(* CODESYS project Revisora(2)_V3_0_2k.project
   Company: Schneider Electric
   Title: Revisora
   Author: Frank Willian
   Version: 2.0.0.0

Project tree, tasks and I/O mapping:
  MyController : TM241CE40T/U, Schneider Electric, order no. TM241CE40T/U, version 4.0.6.18
    application Application
      libraries: SysTime, 3.4.1.20 (System)
      task MAST (cyclic, interval 10 ms, priority 15, watchdog 100 ms x 1) calls R00_main
      task Task1ms (cyclic, interval 1 ms, priority 1) calls RB01_enableReb
      global variables GVL
      01_Maquina/
        program R06_principal [LD]
        program R01_firstScan [LD]
        program R05_comando [LD]
        program R20_acessorios [LD]
        program R99_calcTempos [ST]
        program R00_main [LD]
        program R30_receita [ST]
        program R19_cilindros [LD]
        program R18_alinhador [LD]
        program R50_reset [ST]
      Structs/
        data type _exec_bits
        data type _eixo_drive
        data type _eixo_home
        data type _eixo_auto
        data type _receita
        data type _eixo
      05_IHM/
        program I02_alarmes [ST]
        program I06_textoConfirma [LD]
        program I01_geral [LD]
        program I03_mensagens [ST]
      03_Nip/
        program NP03_auto [LD]
        program NP01_geral [LD]
        program NP06_jog [LD]
        program NP09_sentido [ST]
        program NP04_parada [LD]
        program NP02_enableNip [LD]
        program NP07_veloc [ST]
        program NP20_JogTest [ST]
      global variables PersistentVars
      global variables IHM
      Symbol configuration
      Visu/
      10_Relogio/
        function block GetDateAndTime [CFC]
        function block SetDateAndTime [CFC]
        program AjustaDataHora [LD]
      image pool Imagens
      11_FB/
        function block RTO [ST]
      02_Rebobinadores/
        program RB01_enableReb [LD]
        program RB05_sentido [ST]
        program RB03_analog [LD]
        program RB04_saidas [LD]
      19_Ultra/
        program U10_auto [LD]
    Cartridge_1 : Cartridge, Schneider Electric, version 4.0.6.18
    Cartridge_2 : Cartridge, Schneider Electric, version 4.0.6.18
    IO_Bus : IO bus - TM3, Schneider Electric, version 4.0.6.18
      Saidas_Analog : TM3AQ2/G, Schneider Electric, order no. TM3AQ2/G, version 1.0.0.12
          settings: KPI Configuration.KPI Configuration[0] = 17; KPI Configuration.KPI Configuration[1] = 17; KPI Configuration.KPI Configuration[2] = 240; KPI Configuration.KPI Configuration[3] = 216; KPI Configuration.KPI Configuration[4] = 240; KPI Configuration.KPI Configuration[5] = 216; KPI Configuration.KPI Configuration[6] = 16; KPI Configuration.KPI Configuration[7] = 39; KPI Configuration.KPI Configuration[8] = 16; KPI Configuration.KPI Configuration[9] = 39
          output analoReb01 : INT  // QW0
          output analoReb02 : INT  // QW1
          input  ibAnalog_IBStatusQW0 : BYTE  // IBStatusQW0
          input  ibAnalog_IBStatusQW1 : BYTE  // IBStatusQW1
      Entradas_Analog : TM3AI4/G, Schneider Electric, order no. TM3AI4/G, version 1.0.0.15
          settings: KPI Configuration.KPI Configuration[0] = 34; KPI Configuration.KPI Configuration[1] = 34; KPI Configuration.KPI Configuration[5] = 0; KPI Configuration.KPI Configuration[7] = 0; KPI Configuration.KPI Configuration[12] = 32; KPI Configuration.KPI Configuration[13] = 78; KPI Configuration.KPI Configuration[14] = 32; KPI Configuration.KPI Configuration[15] = 78
          input  ia_sensorUltraSom_1 : INT  // IW0
          input  ia_sensorUltraSom_2 : INT  // IW1
          input  iiModule_1_IW2 : INT  // IW2
          input  iiModule_1_IW3 : INT  // IW3
          input  ibModule_1_IBStatusIW0 : BYTE  // IBStatusIW0
          input  ibModule_1_IBStatusIW1 : BYTE  // IBStatusIW1
          input  ibModule_1_IBStatusIW2 : BYTE  // IBStatusIW2
          input  ibModule_1_IBStatusIW3 : BYTE  // IBStatusIW3
    COM_Bus : COM bus, Schneider Electric, version 4.0.6.18
    Ethernet_1 : Ethernet Network, Schneider Electric, version 4.0.6.18
        settings: IPAddress = [192, 168, 1, 10]; SubnetMask = [255, 255, 255, 0]; WebServer = TRUE; FTP Server = TRUE; SoMachine Protocol = TRUE; Modbus Server = TRUE; NetManage Protocol = TRUE; SNMP protocol = TRUE; WebVisu protocol = TRUE
    Serial_Line_1 : Serial line, Schneider Electric, version 4.0.6.18
      SoMachine_Network_Manager : SoMachine-Network Manager, Schneider Electric, version 4.0.0.2
    Serial_Line_2 : Serial line, Schneider Electric, version 4.0.6.18
      Modbus_Manager : Modbus Manager, Schneider Electric, version 4.0.0.2
    DI : Digital Inputs, Schneider Electric, version 4.0.6.18
        input  i_releEmergencia : BOOL  // IDW0.I0
        input  i_btReset : BOOL  // IDW0.I1
        input  i_ligaRevisora : BOOL  // IDW0.I2
        input  i_sentido : BOOL  // IDW0.I4
        input  i_cortina : BOOL  // IDW0.I6
        input  i_finalDeContagem : BOOL  // IDW0.I9
        unmapped channels: IDW0, IB1
    DQ : Digital Outputs, Schneider Electric, version 4.0.6.18
        settings: Outputs Usage = 15
        output o_enableReb01 : BOOL  // QW0.Q4
        output o_enableNip : BOOL  // QW0.Q5
        output o_enableReb02 : BOOL  // QW0.Q6
        output o_alinhador : BOOL  // QW0.Q7
        output o_mesaCentro : BOOL  // QW0.Q8
        output o_cilindroNip : BOOL  // QW0.Q9
        output o_mesaAuto : BOOL  // QW0.Q10
        output o_abilitaPulsoNip : BOOL  // QW0.Q11
        output qbDQ_QB1 : BYTE  // QB1
        unmapped channels: QW0
    Counters : Counters, Schneider Electric, version 4.0.6.18
    Pulse_Generators : Pulse Generators, Schneider Electric, version 4.0.6.18
        settings: Instance name = 'nip_PTO'; B output History = 'old=-1 new=1'; A output History = 'old=-1 new=0'; Temporary Instance name = 'nip_PTO'; Instance name = 'selag_PTO'; B output History = 'old=-1 new=3'; A output History = 'old=-1 new=2'; Temporary Instance name = 'selag_PTO'
  HMISTU855 : HMIS5T, Schneider Electric, order no. HMIS5T, version 3.5.3.54
    HMI Application
    Ethernet
      SoMachine_Network_Manager2 : SoMachine-Network Manager, Schneider Electric, version 4.0.0.2
    USB
      SoMachine_Network_Manager3 : SoMachine-Network Manager, Schneider Electric, version 4.0.0.2
    COM1
      SoMachine_Network_Manager1 : SoMachine-Network Manager, Schneider Electric, version 4.0.0.2
  6c0f7fb6-600b-4c93-9262-20cdc603757e
  text list GlobalTextList
  5ce3da45-db07-42e7-a21c-a00fff4ed8f6|C:\_Clientes\Opuspac\Doc\Figuras\Botao.png
  5ce3da45-db07-42e7-a21c-a00fff4ed8f6|C:\_Clientes\Opuspac\Doc\Figuras\Botao_ps.png
  5ce3da45-db07-42e7-a21c-a00fff4ed8f6|C:\_Clientes\Opuspac\Doc\Figuras\LogoOpus.jpg
  Vijeo Designer Project Container
*)

// MyController/Application/Structs/_exec_bits
TYPE _exec_bits :
STRUCT
	RQ					: BOOL;
	IP					: BOOL;
	DN					: BOOL;
	Fase				: DINT;
	Mask				: DINT;
END_STRUCT
END_TYPE

// MyController/Application/Structs/_eixo_drive
TYPE _eixo_drive :
STRUCT
	falha			: MC_ReadAxisError_PTO;
	posicao			: MC_ReadActualPosition_PTO;
	power			: MC_Power_PTO;
	reset			: MC_Reset_PTO;
	state			: MC_ReadMotionState_PTO;
	status			: MC_ReadStatus_PTO;
	stop			: MC_Stop_PTO;
END_STRUCT
END_TYPE

// MyController/Application/Structs/_eixo_home
TYPE _eixo_home :
STRUCT
	RQ					: BOOL;
	IP					: BOOL;
	DN					: BOOL;
	Fase				: DINT;
	Mask				: DINT;
	movVeloc			: MC_MoveVelocity_PTO;
	movRelat			: MC_MoveRelative_PTO;
	movStop				: ARRAY[1..2] OF MC_Stop_PTO;
	setPos				: MC_SetPosition_PTO;
END_STRUCT
END_TYPE

// MyController/Application/Structs/_eixo_auto
TYPE _eixo_auto :
STRUCT
	movVeloc					: ARRAY [1..3] OF MC_MoveVelocity_PTO;
	movAbs						: MC_MoveAbsolute_PTO;
	movRelat					: ARRAY [0..3] OF MC_MoveRelative_PTO;
	movStop						: MC_Stop_PTO;
	setPos						: MC_SetPosition_PTO;
END_STRUCT
END_TYPE

// MyController/Application/Structs/_receita
TYPE _receita :
STRUCT
	
	velocDesb		: DINT;
	velocReb		: DINT;
	freioDesb		: INT;
	freioReb		: INT;
	torqueDesb		: INT;
	torqueReb		: INT;

END_STRUCT
END_TYPE

// MyController/Application/Structs/_eixo
TYPE _eixo :
STRUCT
	auto				: _eixo_auto;
	home				: _eixo_home;
	drive				: _eixo_drive;
	falha				: BOOL;
	posicaoAtual		: DINT;
	calcula				: BOOL;
	parando				: BOOL;
	pausa				: BOOL;
	constMove			: BOOL;
	errorStop			: BOOL;
END_STRUCT
END_TYPE

// MyController/Application/GVL
VAR_GLOBAL
	
	jogNip						: BOOL;
	jogRebEsq					: BOOL;
	jogRebDir					: BOOL;
	jogDirecao					: BOOL;
	jogAbilita					: BOOL;
	jogEnebleGeral				: BOOL;
	jogCilindroNip				: BOOL;
	valorPorcRebobinador		: ARRAY [1..2] OF REAL;
	tempoAtrasoAposDesligar		: BOOL;
	troggerTest					: BOOL;
	cortinaOk					: BOOL;
	mudaVeloc					: BOOL;
	auxAnaloReb01				: INT;
	auxAnaloReb02				: INT;
	abilitaTrocaVeloc			: BOOL;
	abilitaPulsoNip				: _exec_bits;
	T_desabilitaPulsoNip		: TON;
	tpoDesabilitaPulsoNip		: BOOL;
	
	
	// transições
	psBtCiclo					: BOOL;

	// Variaveis gerais
	alarmeReset					: BOOL;
	alarmeResetInd				: BOOL;
	alwaysOff					: BOOL;
	alwaysOn					: BOOL;
	calcGeral					: BOOL;
	calcTempos					: BOOL;
	comandoOff					: BOOL;
	emergOk						: BOOL;
	existeAlarme				: BOOL;
	firstScan					: BOOL;
	injecaoTpoOff				: BOOL;
	ladoDir						: BOOL;
	ladoEsq						: BOOL;
	liberaCiclo					: BOOL;
	ligaAlinhador				: BOOL;
	livreComando				: BOOL;
	livreStart					: BOOL;
	ligaMaq						: BOOL;
	manual						: BOOL;
	mesaCentro					: BOOL;
	modoAutomatico				: BOOL;
	nipEmMove					: BOOL;
	nipPausado					: BOOL;
	partidaOK					: BOOL;
	partidaLenta				: BOOL;
	velocPartida				: BOOL;		
	pisca						: BOOL;
	piscaRapido					: BOOL;
	primeiroCiclo				: BOOL;
	start						: BOOL;
	sentidoDesbobinar			: BOOL;
	sentidoRebobinar			: BOOL;
	torqueParada				: BOOL;
	triggerBobina				: BOOL;
	triggerValorDesbReb			: BOOL;
	
	tpoInicio					: TIME;
	
	revisora					: _eixo;
	nip							: _eixo;

	TL_inicializa				: TON;
	T_nipLiga					: TON;
	
	alinhador					: _exec_bits;
	ciclo						: _exec_bits;
	contagem					: _exec_bits;
	cilNip						: _exec_bits;
	comando						: _exec_bits;
	enbReb						: _exec_bits;
	enbNip						: _exec_bits;
	liga						: _exec_bits;
	desliga						: _exec_bits;
	jogNeg						: _exec_bits;
	jogPos						: _exec_bits;
	nipMove						: _exec_bits;
	nipParada					: _exec_bits;
	nipStop						: _exec_bits;
	principal					: _exec_bits;	


	porcRebobinador				: ARRAY [1..2] OF REAL;
	rebobiPorc 					: ARRAY [1..2] OF LIN_TRAFO;
	
    //Sincroniza e ajusta o relógio da IHM
	AnoSet						: UINT;
	ClkScan						: BOOL;
	AjustaHora					: BOOL;
	MesSet						: UINT;
	DiaSet						: UINT;
	HoraSet						: UINT;
	MinutoSet					: UINT;
	SegundoSet					: UINT;
	AnoAtual					: UINT;
	MesAtual					: UINT;
	DiaAtual					: UINT;
	HoraAtual					: UINT;
	MinutoAtual					: UINT;
	SegundoAtual				: UINT;	
	sink						: BOOL;

(*	=================== ALARMES ===================
	Obs: alarme[0]- Não utilizado
*)
	alarme						: ARRAY[0..50] OF BOOL;
	alarmes						: _exec_bits;
	mensagem					: ARRAY[0..50] OF BOOL;
	numAlarme					: SINT;
		
(*	=================== Alterações ===================  *)
	ativoManual					: BOOL;
	tpoArAtivo					: TIME;

(*	=================== Ultrassonico ===================  *)	
	rebobTorqueOper				: ARRAY[0..2] OF REAL;
	desbobTorqueOper			: ARRAY[0..2] OF REAL;
	analogTorqueDrive			: ARRAY[0..2] OF INT;


END_VAR

// MyController/Application/PersistentVars
VAR_GLOBAL PERSISTENT RETAIN
	versaoSoftware				: REAL:= 1.00;
	pi							: REAL:= 3.1415926;
	paramFab					: BOOL:= TRUE;
	numRec						: SINT;
	displayState				: INT;
	jogVelocNip					: DINT;
	revisoraVelocNip			: DINT;
	valorJogRebob01				: INT;
	valorJogRebob02				: INT;
		
	// NIP
	auxVeloc					: ARRAY[0..4] OF BOOL;
	saidaReb					: ARRAY[0..1] OF BOOL;
	M_diamRolo					: DINT:= 34;
	M_revisoraVeloc				: DINT;
	M_revisoraAcel				: DINT:= 800;
	M_revisoraDecel				: DINT:= 200;
	M_pulsosParar				: DINT;
	parseAnalog					: ARRAY[0..1] OF INT;
	ihm_velocidade				: DINT:= 10;
	ihm_tempoInicio				: DINT:= 10;
	visLadoDir					: BOOL;
	visLadoEsq					: BOOL;
	
	veloc						: ARRAY[0..4] OF DINT;
	delayTorq					: ARRAY[0..1] OF TIME;
	sentido						: INT;
	
	bobina			 			: ARRAY[0..5] OF _receita;	
	bobinaAtual					: _receita;
	
	//	========= ultrassonico ===========	
	ihm_btUltraSomHab			: BOOL;
	
	//	========= desbobinador ===========	
	M_desbobTorqueMin				: ARRAY[0..2] OF REAL;
	M_desbobTorqueMax				: ARRAY[0..2] OF REAL;
	M_desbobTorqueOper				: ARRAY[0..2] OF REAL;
	valorDesbobTorqueMin			: REAL;
	valorDesbobTorqueMax			: REAL;
	
	//  ========== Rebobinador ===========
	M_rebobTorqueMin				: ARRAY[0..2] OF REAL;
	M_rebobTorqueMax				: ARRAY[0..2] OF REAL;
	M_rebobTorqueOper				: ARRAY[0..2] OF REAL;
	valorRebobTorqueMin				: REAL;
	valorRebobTorqueMax				: REAL;

END_VAR

// MyController/Application/IHM
VAR_GLOBAL
	ihm_alarme					: ARRAY[0..50] OF BOOL;
	ihm_alarmeReset				: BOOL;
	ihm_alarmeResetInd			: BOOL;
	ihm_bannerConfirma			: BOOL;
	ihm_bannerMensagem			: BOOL;
	ihm_confirmaV				: BOOL;
	ihm_confirmaX				: BOOL;
	ihm_mensagem				: DINT;
	ihm_numReceita				: SINT;
	ihm_telaHome				: BOOL;
	ihm_telaAtual				: INT;
	ihm_textoConfirma			: DINT;
	ihm_textoProced				: DINT;
	ihm_velocMedida				: DINT;
	ihm_inverte					: BOOL;
	ihm_cilindroNip				: BOOL;
	ihm_alinhador				: BOOL;
	nome						: WSTRING;
	
	ihm_valorDesb				: ARRAY[0..2] OF REAL;
	ihm_valorReb				: ARRAY[0..2] OF REAL;
	
	ihm_desbobInc				: BOOL;
	ihm_desbobDec				: BOOL;
	
	ihm_rebobInc				: BOOL;
	ihm_rebobDec				: BOOL;

END_VAR

// MyController/Application/01_Maquina/R00_main
PROGRAM R00_main
VAR
END_VAR

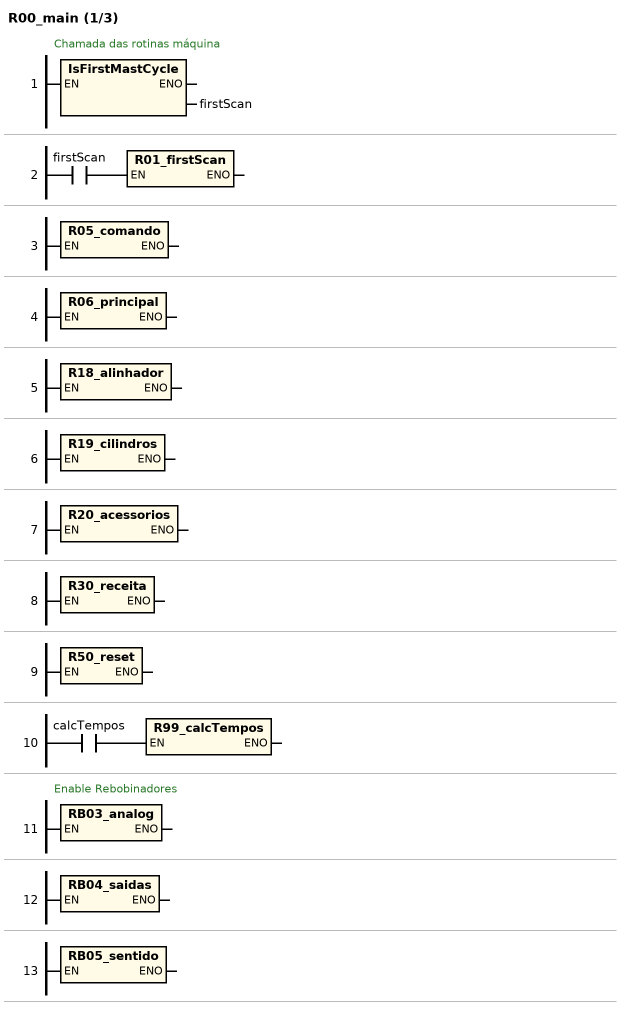
// NETWORK 1
// Chamada das rotinas máquina
firstScan := IsFirstMastCycle();

// NETWORK 2
IF firstScan THEN R01_firstScan(); END_IF

// NETWORK 3
R05_comando();

// NETWORK 4
R06_principal();

// NETWORK 5
R18_alinhador();

// NETWORK 6
R19_cilindros();

// NETWORK 7
R20_acessorios();

// NETWORK 8
R30_receita();

// NETWORK 9
R50_reset();

// NETWORK 10
IF calcTempos THEN R99_calcTempos(); END_IF

// NETWORK 11
// Enable Rebobinadores
RB03_analog();

// NETWORK 12
RB04_saidas();

// NETWORK 13
RB05_sentido();

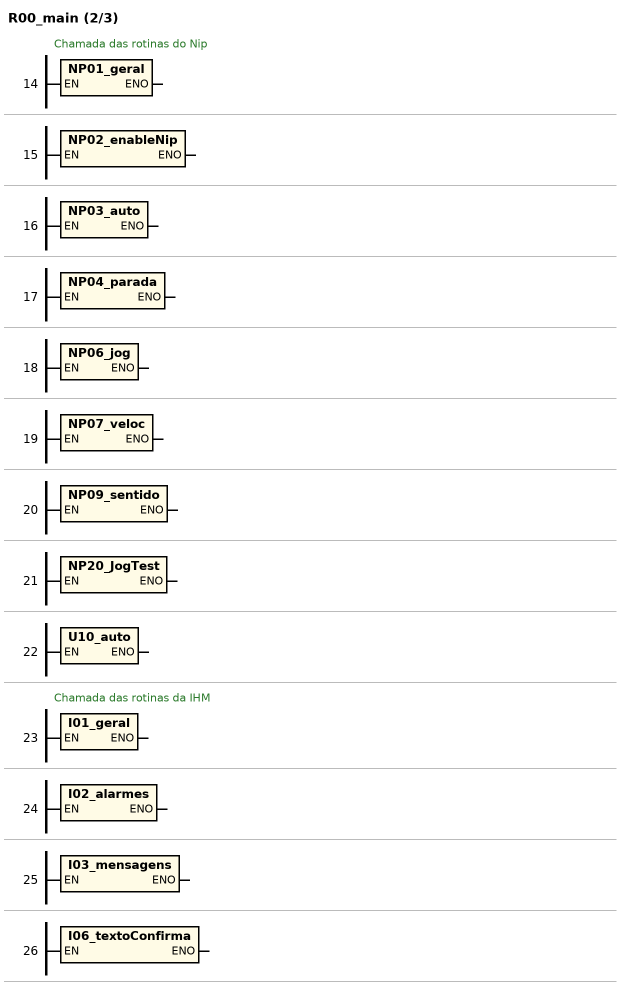
// NETWORK 14
// Chamada das rotinas do Nip
NP01_geral();

// NETWORK 15
NP02_enableNip();

// NETWORK 16
NP03_auto();

// NETWORK 17
NP04_parada();

// NETWORK 18
NP06_jog();

// NETWORK 19
NP07_veloc();

// NETWORK 20
NP09_sentido();

// NETWORK 21
NP20_JogTest();

// NETWORK 22
U10_auto();

// NETWORK 23
// Chamada das rotinas da IHM
I01_geral();

// NETWORK 24
I02_alarmes();

// NETWORK 25
I03_mensagens();

// NETWORK 26
I06_textoConfirma();

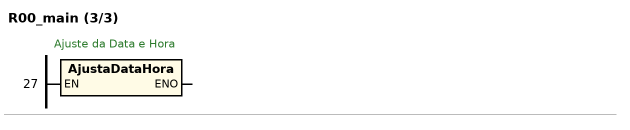
// NETWORK 27
// Ajuste da Data e Hora
AjustaDataHora();

END_PROGRAM

// MyController/Application/01_Maquina/R01_firstScan
PROGRAM R01_firstScan
VAR
END_VAR

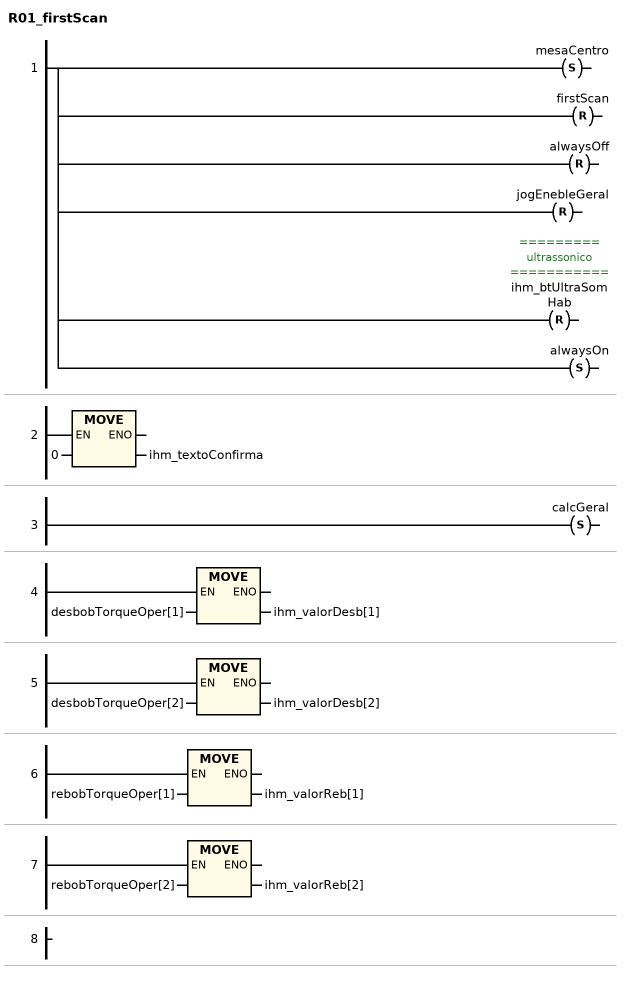
// NETWORK 1
//   ihm_btUltraSomHab: ========= ultrassonico ===========
mesaCentro S= TRUE;
firstScan R= TRUE;
alwaysOff R= TRUE;
jogEnebleGeral R= TRUE;
ihm_btUltraSomHab R= TRUE;
alwaysOn S= TRUE;

// NETWORK 2
ihm_textoConfirma := 0;

// NETWORK 3
calcGeral S= TRUE;

// NETWORK 4
ihm_valorDesb[1] := desbobTorqueOper[1];

// NETWORK 5
ihm_valorDesb[2] := desbobTorqueOper[2];

// NETWORK 6
//   rebobTorqueOper[1]: =================== Ultrassonico ===================
ihm_valorReb[1] := rebobTorqueOper[1];

// NETWORK 7
//   rebobTorqueOper[2]: =================== Ultrassonico ===================
ihm_valorReb[2] := rebobTorqueOper[2];

// NETWORK 8

END_PROGRAM

// MyController/Application/01_Maquina/R05_comando
PROGRAM R05_comando
VAR
	TL_comando				: TON;
END_VAR
VAR // added by the converter: edge detectors and wires of the graphical bodies
    _rt1 : R_TRIG;
    _ft1, _ft2 : F_TRIG;
    _w1 : BOOL;
END_VAR

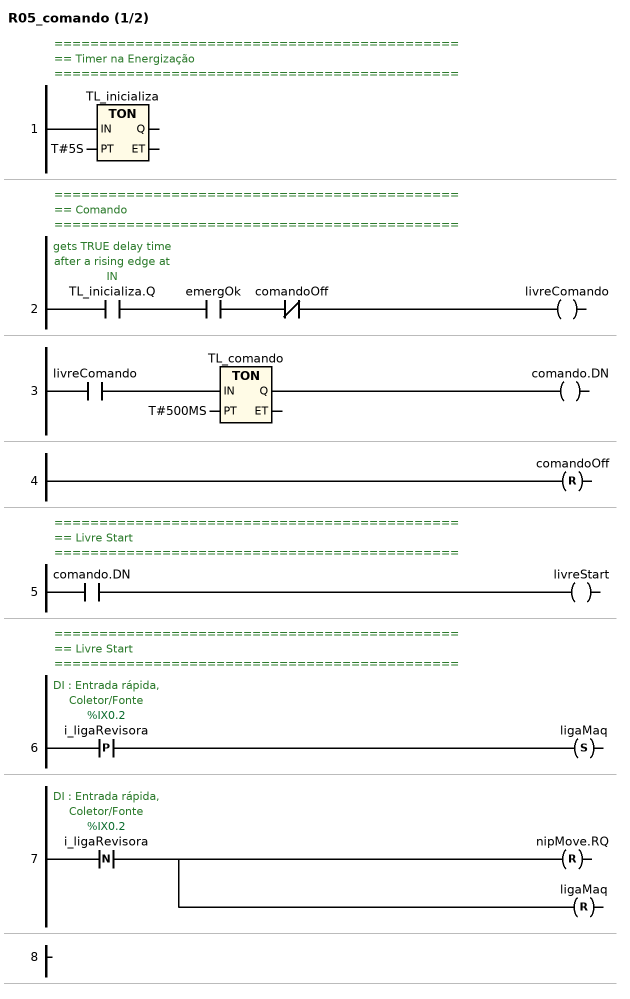
// NETWORK 1
// =============================================
// == Timer na Energização
// =============================================
TL_inicializa(IN := TRUE, PT := T#5S); // TON

// NETWORK 2
// =============================================
// == Comando
// =============================================
//   TL_inicializa.Q: gets TRUE delay time after a rising edge at IN
livreComando := TL_inicializa.Q AND emergOk AND NOT comandoOff;

// NETWORK 3
TL_comando(IN := livreComando, PT := T#500MS); // TON
comando.DN := TL_comando.Q;

// NETWORK 4
comandoOff R= TRUE;

// NETWORK 5
// =============================================
// == Livre Start
// =============================================
livreStart := comando.DN;

// NETWORK 6
// =============================================
// == Livre Start
// =============================================
//   i_ligaRevisora: DI : Entrada rápida, Coletor/Fonte | AT %IX0.2
_rt1(CLK := i_ligaRevisora);
ligaMaq S= _rt1.Q;

// NETWORK 7
//   i_ligaRevisora: DI : Entrada rápida, Coletor/Fonte | AT %IX0.2
_ft1(CLK := i_ligaRevisora);
nipMove.RQ R= _ft1.Q;
ligaMaq R= _ft1.Q;

// NETWORK 8

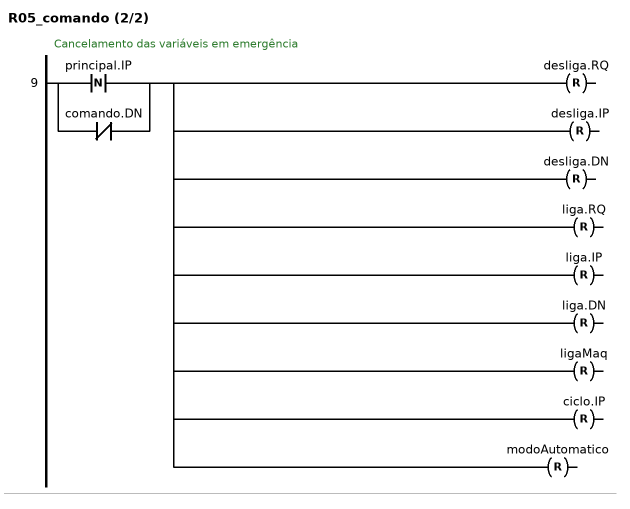
// NETWORK 9
// Cancelamento das variáveis em emergência
_ft2(CLK := principal.IP);
_w1 := _ft2.Q OR NOT comando.DN;
desliga.RQ R= _w1;
desliga.IP R= _w1;
desliga.DN R= _w1;
liga.RQ R= _w1;
liga.IP R= _w1;
liga.DN R= _w1;
ligaMaq R= _w1;
ciclo.IP R= _w1;
modoAutomatico R= _w1;

END_PROGRAM

// MyController/Application/01_Maquina/R06_principal
PROGRAM R06_principal
VAR

	T_inicio				: ARRAY[0..2] OF TON;
	T_partida				: TON;
	T_parada				: TON;
	T_delayMudaVeloc: TON;
	T_delay: TON;
END_VAR
VAR // added by the converter: edge detectors and wires of the graphical bodies
    _w1, _w2, _w3, _w4 : BOOL;
    _ft1 : F_TRIG;
END_VAR

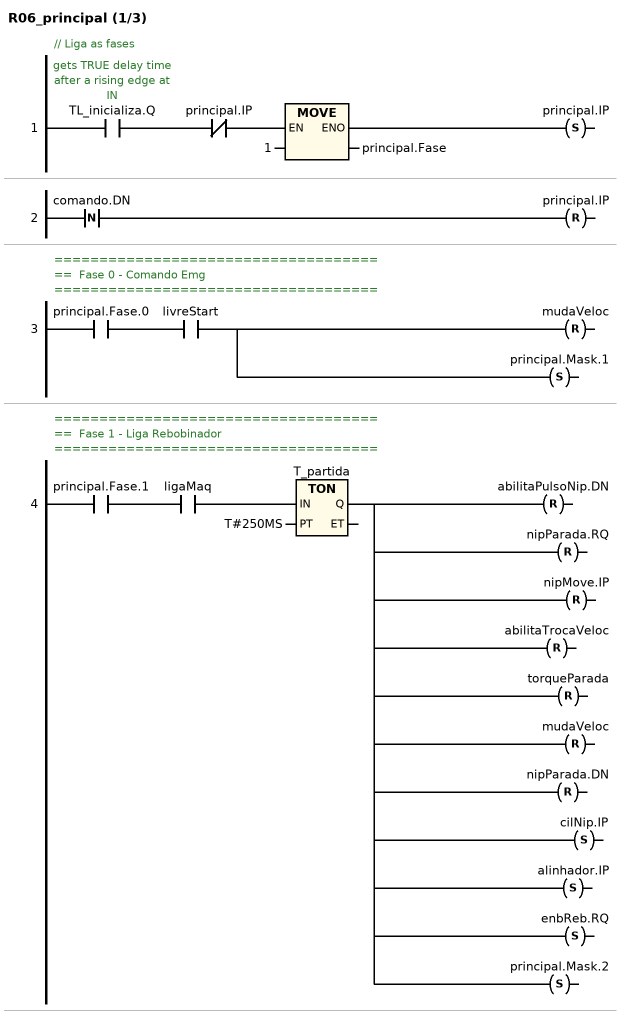
// NETWORK 1
// // Liga as fases
//   TL_inicializa.Q: gets TRUE delay time after a rising edge at IN
_w1 := TL_inicializa.Q AND NOT principal.IP;
IF _w1 THEN principal.Fase := 1; END_IF
principal.IP S= _w1;

// NETWORK 2
_ft1(CLK := comando.DN);
principal.IP R= _ft1.Q;

// NETWORK 3
// ====================================
// ==  Fase 0 - Comando Emg
// ====================================
_w2 := principal.Fase.0 AND livreStart;
mudaVeloc R= _w2;
principal.Mask.1 S= _w2;

// NETWORK 4
// ====================================
// ==  Fase 1 - Liga Rebobinador
// ====================================
T_partida(IN := principal.Fase.1 AND ligaMaq, PT := T#250MS); // TON
abilitaPulsoNip.DN R= T_partida.Q;
nipParada.RQ R= T_partida.Q;
nipMove.IP R= T_partida.Q;
abilitaTrocaVeloc R= T_partida.Q;
torqueParada R= T_partida.Q;
mudaVeloc R= T_partida.Q;
nipParada.DN R= T_partida.Q;
cilNip.IP S= T_partida.Q;
alinhador.IP S= T_partida.Q;
enbReb.RQ S= T_partida.Q;
principal.Mask.2 S= T_partida.Q;

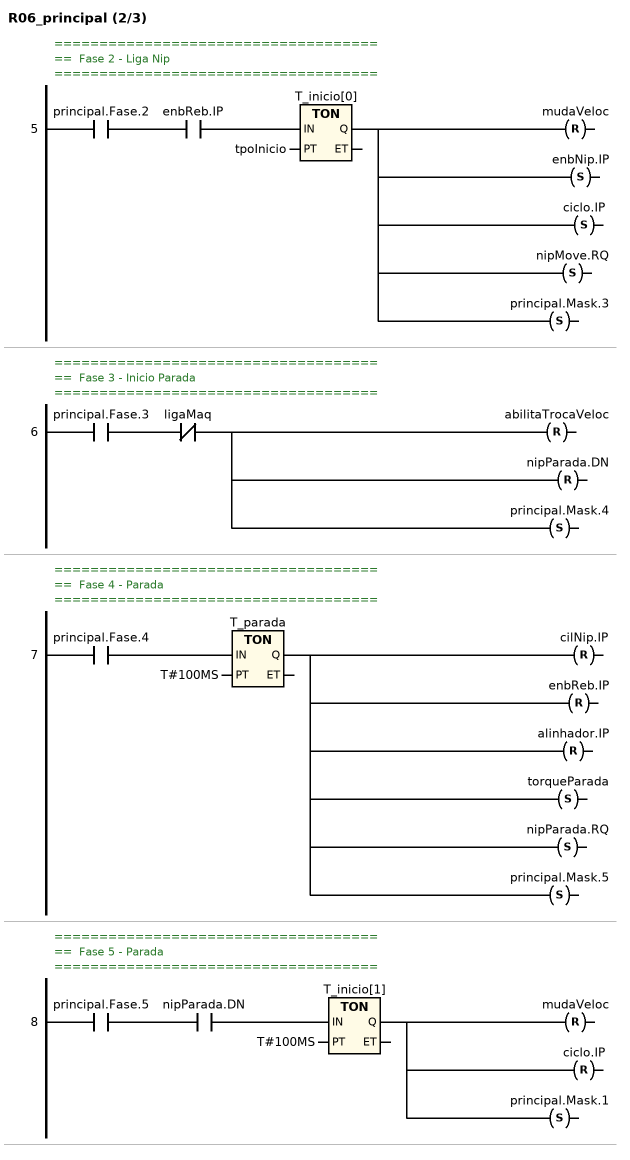
// NETWORK 5
// ====================================
// ==  Fase 2 - Liga Nip
// ====================================
T_inicio[0](IN := principal.Fase.2 AND enbReb.IP, PT := tpoInicio); // TON
mudaVeloc R= T_inicio[0].Q;
enbNip.IP S= T_inicio[0].Q;
ciclo.IP S= T_inicio[0].Q;
nipMove.RQ S= T_inicio[0].Q;
principal.Mask.3 S= T_inicio[0].Q;

// NETWORK 6
// ====================================
// ==  Fase 3 - Inicio Parada
// ====================================
_w3 := principal.Fase.3 AND NOT ligaMaq;
abilitaTrocaVeloc R= _w3;
nipParada.DN R= _w3;
principal.Mask.4 S= _w3;

// NETWORK 7
// ====================================
// ==  Fase 4 - Parada
// ====================================
T_parada(IN := principal.Fase.4, PT := T#100MS); // TON
cilNip.IP R= T_parada.Q;
enbReb.IP R= T_parada.Q;
alinhador.IP R= T_parada.Q;
torqueParada S= T_parada.Q;
nipParada.RQ S= T_parada.Q;
principal.Mask.5 S= T_parada.Q;

// NETWORK 8
// ====================================
// ==  Fase 5 - Parada
// ====================================
T_inicio[1](IN := principal.Fase.5 AND nipParada.DN, PT := T#100MS); // TON
mudaVeloc R= T_inicio[1].Q;
ciclo.IP R= T_inicio[1].Q;
principal.Mask.1 S= T_inicio[1].Q;

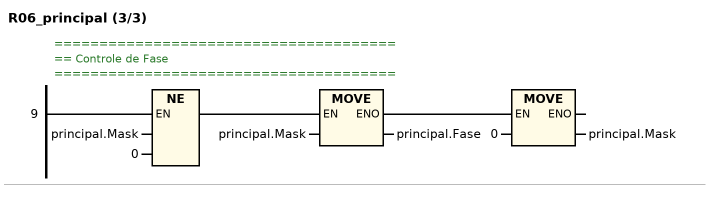
// NETWORK 9
// ======================================
// == Controle de Fase
// ======================================
_w4 := principal.Mask <> 0;
IF _w4 THEN principal.Fase := principal.Mask; END_IF
IF _w4 THEN principal.Mask := 0; END_IF

END_PROGRAM

// MyController/Application/01_Maquina/R18_alinhador
PROGRAM R18_alinhador
VAR
	T_MesaCentro: ARRAY[0..1] OF TON;
	mesaCentro: BOOL;
END_VAR
VAR // added by the converter: edge detectors and wires of the graphical bodies
    _rt1 : R_TRIG;
    _ft1 : F_TRIG;
END_VAR

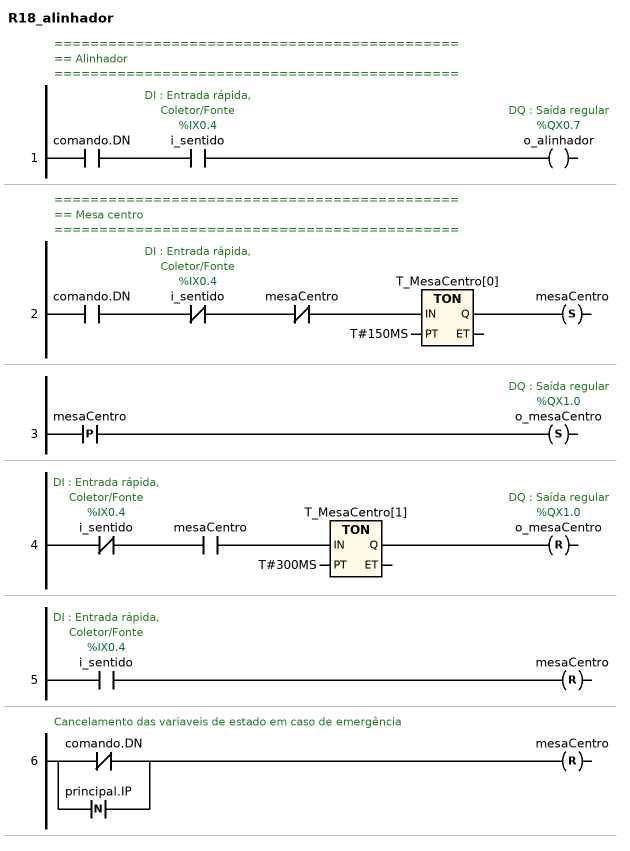
// NETWORK 1
// =============================================
// == Alinhador
// =============================================
//   i_sentido: DI : Entrada rápida, Coletor/Fonte | AT %IX0.4
//   o_alinhador: DQ : Saída regular | AT %QX0.7
o_alinhador := comando.DN AND i_sentido;

// NETWORK 2
// =============================================
// == Mesa centro
// =============================================
//   i_sentido: DI : Entrada rápida, Coletor/Fonte | AT %IX0.4
T_MesaCentro[0](IN := comando.DN AND NOT i_sentido AND NOT mesaCentro, PT := T#150MS); // TON
mesaCentro S= T_MesaCentro[0].Q;

// NETWORK 3
//   o_mesaCentro: DQ : Saída regular | AT %QX1.0
_rt1(CLK := mesaCentro);
o_mesaCentro S= _rt1.Q;

// NETWORK 4
//   i_sentido: DI : Entrada rápida, Coletor/Fonte | AT %IX0.4
//   o_mesaCentro: DQ : Saída regular | AT %QX1.0
T_MesaCentro[1](IN := NOT i_sentido AND mesaCentro, PT := T#300MS); // TON
o_mesaCentro R= T_MesaCentro[1].Q;

// NETWORK 5
//   i_sentido: DI : Entrada rápida, Coletor/Fonte | AT %IX0.4
mesaCentro R= i_sentido;

// NETWORK 6
// Cancelamento das variaveis de estado em caso de emergência
_ft1(CLK := principal.IP);
mesaCentro R= NOT comando.DN OR _ft1.Q;

END_PROGRAM

// MyController/Application/01_Maquina/R19_cilindros
PROGRAM R19_cilindros
VAR
END_VAR
VAR // added by the converter: edge detectors and wires of the graphical bodies
    _ft1 : F_TRIG;
    _w1 : BOOL;
END_VAR

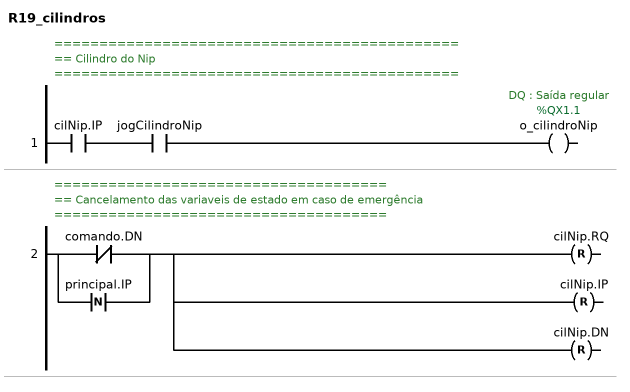
// NETWORK 1
// =============================================
// == Cilindro do Nip
// =============================================
//   o_cilindroNip: DQ : Saída regular | AT %QX1.1
o_cilindroNip := cilNip.IP AND jogCilindroNip;

// NETWORK 2
// =====================================
// == Cancelamento das variaveis de estado em caso de emergência
// =====================================
_ft1(CLK := principal.IP);
_w1 := NOT comando.DN OR _ft1.Q;
cilNip.RQ R= _w1;
cilNip.IP R= _w1;
cilNip.DN R= _w1;

END_PROGRAM

// MyController/Application/01_Maquina/R20_acessorios
PROGRAM R20_acessorios
VAR

	TL_pisca					: BLINK;
	TL_piscaRapido				: BLINK;
	T_atrasoStopNip				: TON;

END_VAR
VAR // added by the converter: edge detectors and wires of the graphical bodies
    _w1, _w2 : BOOL;
END_VAR

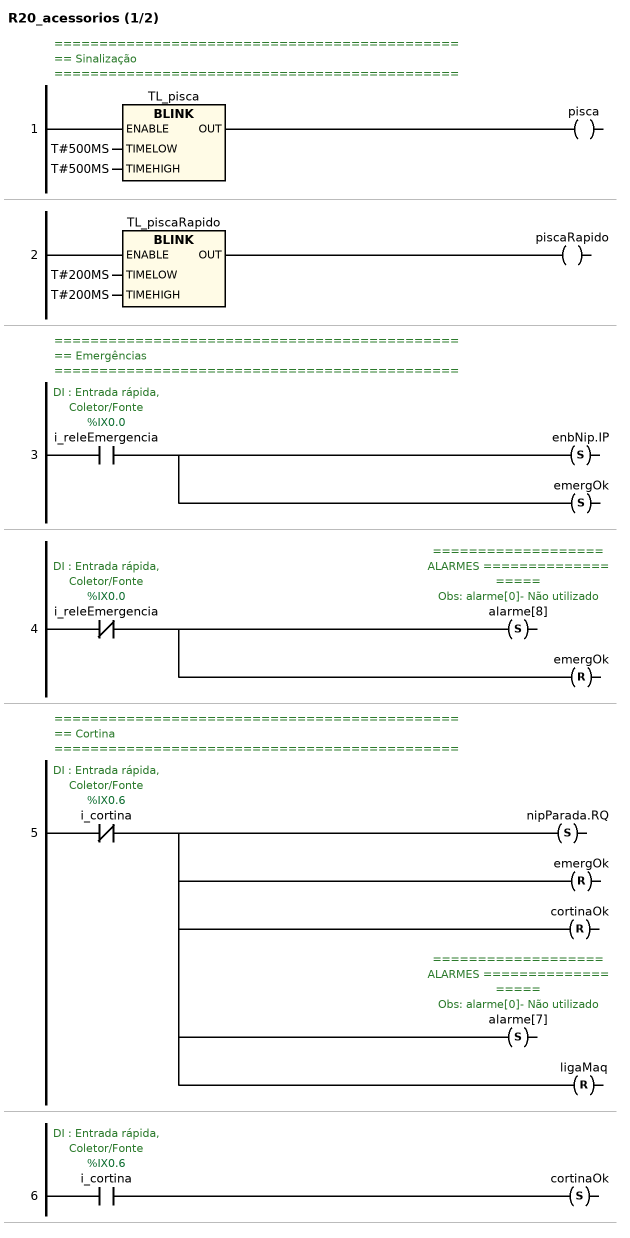
// NETWORK 1
// =============================================
// == Sinalização
// =============================================
TL_pisca(ENABLE := TRUE, TIMELOW := T#500MS, TIMEHIGH := T#500MS); // BLINK
pisca := TL_pisca.OUT;

// NETWORK 2
TL_piscaRapido(ENABLE := TRUE, TIMELOW := T#200MS, TIMEHIGH := T#200MS); // BLINK
piscaRapido := TL_piscaRapido.OUT;

// NETWORK 3
// =============================================
// == Emergências
// =============================================
//   i_releEmergencia: DI : Entrada rápida, Coletor/Fonte | AT %IX0.0
enbNip.IP S= i_releEmergencia;
emergOk S= i_releEmergencia;

// NETWORK 4
//   i_releEmergencia: DI : Entrada rápida, Coletor/Fonte | AT %IX0.0
//   alarme[8]: =================== ALARMES =================== Obs: alarme[0]- Não utilizado
_w1 := NOT i_releEmergencia;
alarme[8] S= _w1;
emergOk R= _w1;

// NETWORK 5
// =============================================
// == Cortina
// =============================================
//   i_cortina: DI : Entrada rápida, Coletor/Fonte | AT %IX0.6
//   alarme[7]: =================== ALARMES =================== Obs: alarme[0]- Não utilizado
_w2 := NOT i_cortina;
nipParada.RQ S= _w2;
emergOk R= _w2;
cortinaOk R= _w2;
alarme[7] S= _w2;
ligaMaq R= _w2;

// NETWORK 6
//   i_cortina: DI : Entrada rápida, Coletor/Fonte | AT %IX0.6
cortinaOk S= i_cortina;
